(* Logix 5000 project; controller FV vendor 1 type 14 code 217 rev 31.11; software revision 31.00; part 29 of 63 *)
(* tags used below, declared in another part *)
   Alarm_Reset : BOOL;
   Default_Check_Time : DINT;
   FR_FV30_AV01 : PlantItem;   // FV30_AV01
   FR_FV30_AV01_ALARM : ALARM_DIGITAL;
   FR_FV30_AV01_C : ALIAS FOR RIO_Rack_2:10:I.Data.4;
   FR_FV30_AV01_O : ALIAS FOR RIO_Rack_2:10:I.Data.0;
   FR_FV30_AV01_RDR : ALIAS FOR RIO_Rack_2:11:O.Data.0;
   FR_FV30_AV04 : PlantItem;   // FV30_AV04
   FR_FV30_AV04_ALARM : ALARM_DIGITAL;
   FR_FV30_AV04_C : ALIAS FOR RIO_Rack_2:10:I.Data.5;
   FR_FV30_AV04_DR : ALIAS FOR RIO_Rack_2:11:O.Data.1;
   FR_FV30_AV04_O : ALIAS FOR RIO_Rack_2:10:I.Data.1;
   FR_FV30_AV05 : PlantItem;   // FV30_AV05
   FR_FV30_AV05_ALARM : ALARM_DIGITAL;
   FR_FV30_AV05_C : ALIAS FOR RIO_Rack_2:10:I.Data.6;
   FR_FV30_AV05_DR : ALIAS FOR RIO_Rack_2:11:O.Data.2;
   FR_FV30_AV05_O : ALIAS FOR RIO_Rack_2:10:I.Data.2;
   FR_FV30_AV06 : PlantItem;   // FV30_AV06
   FR_FV30_AV06_ALARM : ALARM_DIGITAL;
   FR_FV30_AV06_C : ALIAS FOR RIO_Rack_2:10:I.Data.7;
   FR_FV30_AV06_DR : ALIAS FOR RIO_Rack_2:11:O.Data.3;
   FR_FV30_AV06_O : ALIAS FOR RIO_Rack_2:10:I.Data.3;
   FR_FV30_AV07 : PlantItem;   // FV30_AV07
   FR_FV30_AV07_ALARM : ALARM_DIGITAL;
   FR_FV30_AV07_C : ALIAS FOR RIO_Rack_2:10:I.Data.12;
   FR_FV30_AV07_DR : ALIAS FOR RIO_Rack_2:11:O.Data.4;
   FR_FV30_AV07_O : ALIAS FOR RIO_Rack_2:10:I.Data.8;
   FR_VB4_AV04 : PlantItem;   // VB4_AV04
   FR_VB4_AV04_ALARM : ALARM_DIGITAL;
   FR_VB4_AV04_C : ALIAS FOR RIO_Rack_2:7:I.Data.29;
   FR_VB4_AV04_DR : ALIAS FOR RIO_Rack_2:8:O.Data.13;
   FR_VB4_AV04_O : ALIAS FOR RIO_Rack_2:7:I.Data.25;
   FR_VB4_AV05 : PlantItem;   // VB4_AV05
   FR_VB4_AV05_ALARM : ALARM_DIGITAL;
   FR_VB4_AV05_C : ALIAS FOR RIO_Rack_2:7:I.Data.30;
   FR_VB4_AV05_DR : ALIAS FOR RIO_Rack_2:8:O.Data.14;
   FR_VB4_AV05_O : ALIAS FOR RIO_Rack_2:7:I.Data.26;
   FR_VB4_AV06 : PlantItem;   // VB4_AV06
   FR_VB4_AV06_ALARM : ALARM_DIGITAL;
   FR_VB4_AV06_C : ALIAS FOR RIO_Rack_2:7:I.Data.31;
   FR_VB4_AV06_DR : ALIAS FOR RIO_Rack_2:8:O.Data.15;
   FR_VB4_AV06_O : ALIAS FOR RIO_Rack_2:7:I.Data.27;
   FR_VB4_AV07 : PlantItem;   // VB4_AV07
   FR_VB4_AV07_ALARM : ALARM_DIGITAL;
   FR_VB4_AV07_C : ALIAS FOR RIO_Rack_2:9:I.Data.4;
   FR_VB4_AV07_DR : ALIAS FOR RIO_Rack_2:8:O.Data.16;
   FR_VB4_AV07_O : ALIAS FOR RIO_Rack_2:9:I.Data.0;
   FR_VB4_AV08 : PlantItem;   // VB4_AV08
   FR_VB4_AV08_ALARM : ALARM_DIGITAL;
   FR_VB4_AV08_C : ALIAS FOR RIO_Rack_2:9:I.Data.5;
   FR_VB4_AV08_DR : ALIAS FOR RIO_Rack_2:8:O.Data.17;
   FR_VB4_AV08_O : ALIAS FOR RIO_Rack_2:9:I.Data.1;
   FR_VB4_AV09 : PlantItem;   // VB4_AV09
   FR_VB4_AV09_ALARM : ALARM_DIGITAL;
   FR_VB4_AV09_C : ALIAS FOR RIO_Rack_2:9:I.Data.6;
   FR_VB4_AV09_DR : ALIAS FOR RIO_Rack_2:8:O.Data.18;
   FR_VB4_AV09_O : ALIAS FOR RIO_Rack_2:9:I.Data.2;
   FR_VB4_AV10 : PlantItem;   // VB4_AV10
   FR_VB4_AV10_ALARM : ALARM_DIGITAL;
   FR_VB4_AV10_C : ALIAS FOR RIO_Rack_2:9:I.Data.7;
   FR_VB4_AV10_DR : ALIAS FOR RIO_Rack_2:8:O.Data.19;
   FR_VB4_AV10_O : ALIAS FOR RIO_Rack_2:9:I.Data.3;
   FR_VB4_AV11 : PlantItem;   // VB4_AV11
   FR_VB4_AV11_ALARM : ALARM_DIGITAL;
   FR_VB4_AV11_C : ALIAS FOR RIO_Rack_2:9:I.Data.12;
   FR_VB4_AV11_DR : ALIAS FOR RIO_Rack_2:8:O.Data.20;
   FR_VB4_AV11_O : ALIAS FOR RIO_Rack_2:9:I.Data.8;
   FR_VB4_AV12 : PlantItem;   // VB4_AV12
   FR_VB4_AV12_ALARM : ALARM_DIGITAL;
   FR_VB4_AV12_C : ALIAS FOR RIO_Rack_2:9:I.Data.13;
   FR_VB4_AV12_DR : ALIAS FOR RIO_Rack_2:8:O.Data.21;
   FR_VB4_AV12_O : ALIAS FOR RIO_Rack_2:9:I.Data.9;
   FR_VB4_AV13 : PlantItem;   // VB4_AV13
   FR_VB4_AV13_ALARM : ALARM_DIGITAL;
   FR_VB4_AV13_C : ALIAS FOR RIO_Rack_2:9:I.Data.14;
   FR_VB4_AV13_DR : ALIAS FOR RIO_Rack_2:8:O.Data.22;
   FR_VB4_AV13_O : ALIAS FOR RIO_Rack_2:9:I.Data.10;
   FR_VB4_AV14 : PlantItem;   // VB4_AV14
   FR_VB4_AV14_ALARM : ALARM_DIGITAL;
   FR_VB4_AV14_C : ALIAS FOR RIO_Rack_2:9:I.Data.15;
   FR_VB4_AV14_DR : ALIAS FOR RIO_Rack_2:8:O.Data.23;
   FR_VB4_AV14_O : ALIAS FOR RIO_Rack_2:9:I.Data.11;
   FR_VB4_AV15 : PlantItem;   // VB4_AV15
   FR_VB4_AV15_ALARM : ALARM_DIGITAL;
   FR_VB4_AV15_C : ALIAS FOR RIO_Rack_2:9:I.Data.20;
   FR_VB4_AV15_DR : ALIAS FOR RIO_Rack_2:8:O.Data.24;
   FR_VB4_AV15_O : ALIAS FOR RIO_Rack_2:9:I.Data.16;
   FR_VB4_AV17 : PlantItem;   // VB4_AV17
   FR_VB4_AV17_ALARM : ALARM_DIGITAL;
   FR_VB4_AV17_C : ALIAS FOR RIO_Rack_2:9:I.Data.22;
   FR_VB4_AV17_DR : ALIAS FOR RIO_Rack_2:8:O.Data.26;
   FR_VB4_AV17_O : ALIAS FOR RIO_Rack_2:9:I.Data.18;
   FR_VB4_AV18 : PlantItem;   // VB4_AV18
   FR_VB4_AV18_ALARM : ALARM_DIGITAL;
   FR_VB4_AV18_C : ALIAS FOR RIO_Rack_2:9:I.Data.23;
   FR_VB4_AV18_DR : ALIAS FOR RIO_Rack_2:8:O.Data.27;
   FR_VB4_AV18_O : ALIAS FOR RIO_Rack_2:9:I.Data.19;
   FR_VB4_AV19 : PlantItem;   // VB4_AV19
   FR_VB4_AV19_ALARM : ALARM_DIGITAL;
   FR_VB4_AV19_C : ALIAS FOR RIO_Rack_2:9:I.Data.28;
   FR_VB4_AV19_DR : ALIAS FOR RIO_Rack_2:8:O.Data.28;
   FR_VB4_AV19_O : ALIAS FOR RIO_Rack_2:9:I.Data.24;
   FR_VB4_AV20 : PlantItem;   // VB4_AV20
   FR_VB4_AV20_ALARM : ALARM_DIGITAL;
   FR_VB4_AV20_C : ALIAS FOR RIO_Rack_2:9:I.Data.29;
   FR_VB4_AV20_DR : ALIAS FOR RIO_Rack_2:8:O.Data.29;
   FR_VB4_AV20_O : ALIAS FOR RIO_Rack_2:9:I.Data.25;
   FR_VB4_AV21 : PlantItem;   // VB4_AV21
   FR_VB4_AV21_ALARM : ALARM_DIGITAL;
   FR_VB4_AV21_C : ALIAS FOR RIO_Rack_2:9:I.Data.30;
   FR_VB4_AV21_DR : ALIAS FOR RIO_Rack_2:8:O.Data.30;
   FR_VB4_AV21_O : ALIAS FOR RIO_Rack_2:9:I.Data.26;
   FR_VB4_AV22 : PlantItem;   // VB4_AV22
   FR_VB4_AV22_ALARM : ALARM_DIGITAL;
   FR_VB4_AV22_C : ALIAS FOR RIO_Rack_2:9:I.Data.31;
   FR_VB4_AV22_DR : ALIAS FOR RIO_Rack_2:8:O.Data.31;
   FR_VB4_AV22_O : ALIAS FOR RIO_Rack_2:9:I.Data.27;
   FR_VB4_AV23 : PlantItem;   // VB4_AV23
   FR_VB4_AV23_ALARM : ALARM_DIGITAL;
   FR_VB4_AV23_C : ALIAS FOR RIO_Rack_2:9:I.Data.21;
   FR_VB4_AV23_DR : ALIAS FOR RIO_Rack_2:8:O.Data.25;
   FR_VB4_AV23_O : ALIAS FOR RIO_Rack_2:9:I.Data.17;
   Item_Faults_Are_Latched : BOOL;
   Item_Simulation_Flag : BOOL;
   One_Second_One_Scan : ALIAS FOR One_Second_1_scan;
(* FR_Common, continued *)

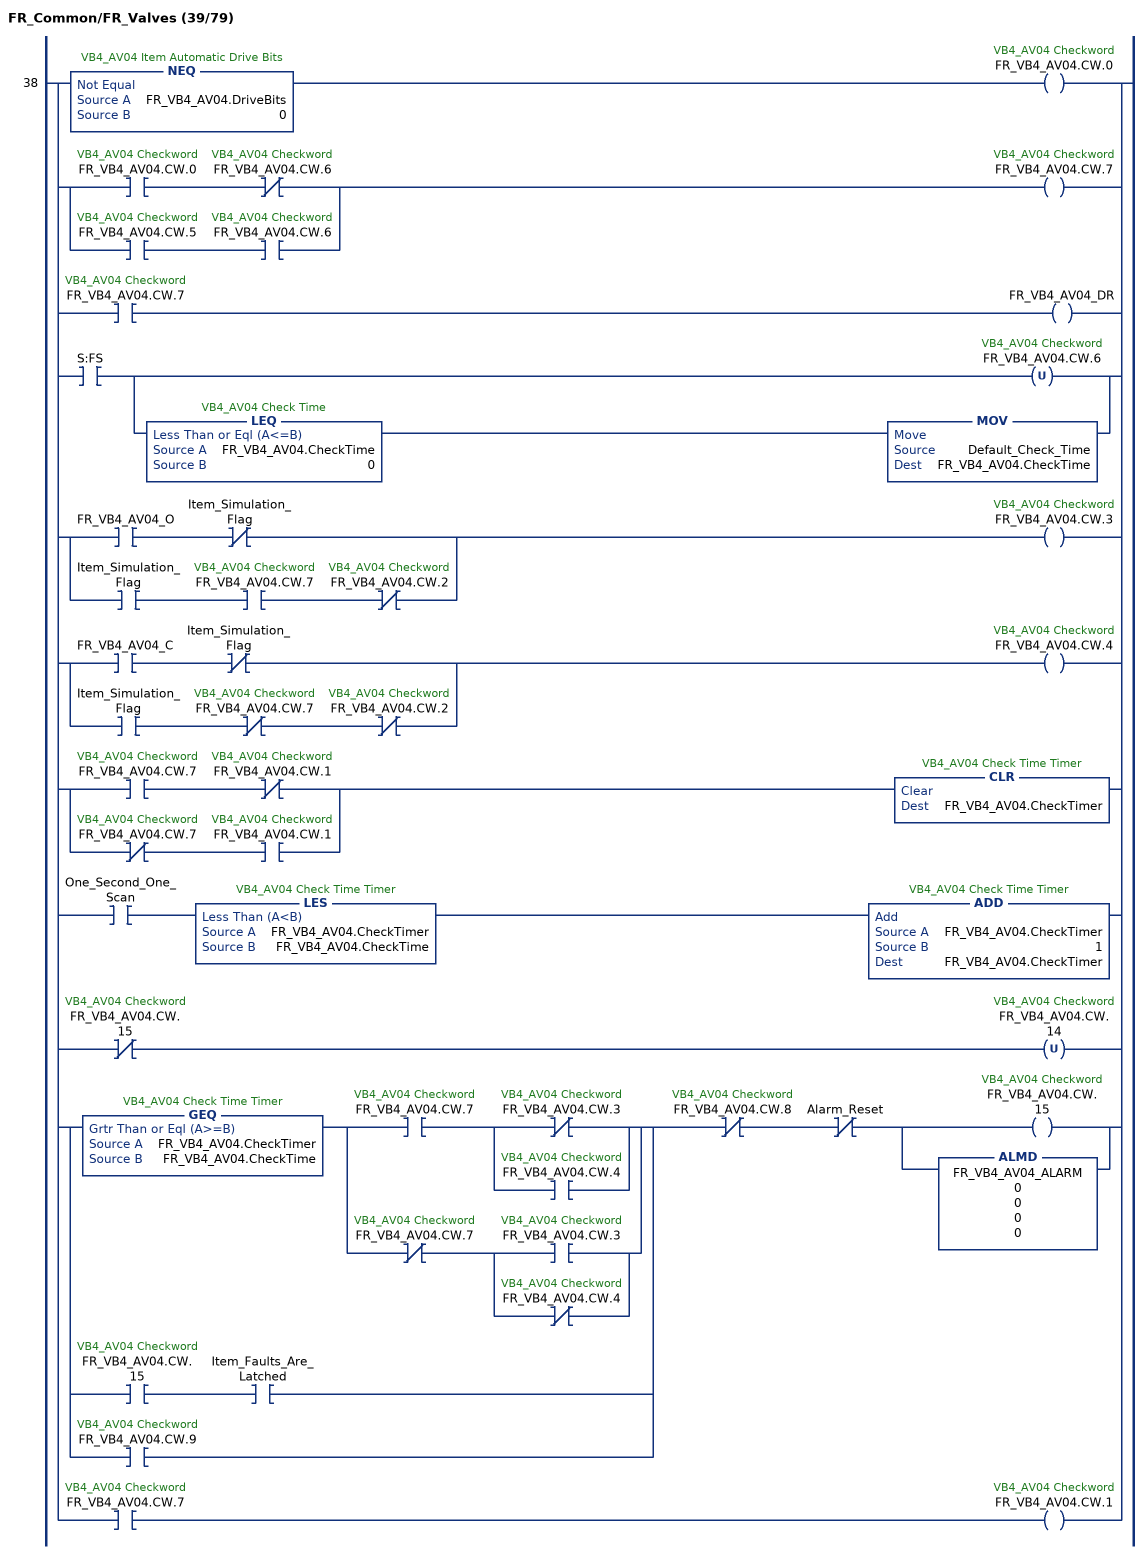
   [picture p592: FR_Common/FR_Valves rungs 38-38]
   38: [NEQ(FR_VB4_AV04.DriveBits,0) OTE(FR_VB4_AV04.CW.0) ,[XIC(FR_VB4_AV04.CW.0) XIO(FR_VB4_AV04.CW.6) ,XIC(FR_VB4_AV04.CW.5) XIC(FR_VB4_AV04.CW.6) ] OTE(FR_VB4_AV04.CW.7) ,XIC(FR_VB4_AV04.CW.7) OTE(FR_VB4_AV04_DR) ,XIC(S:FS) [OTU(FR_VB4_AV04.CW.6) ,LEQ(FR_VB4_AV04.CheckTime,0) MOV(Default_Check_Time,FR_VB4_AV04.CheckTime) ] ,[[XIC(FR_VB4_AV04_O) XIO(Item_Simulation_Flag) ,XIC(Item_Simulation_Flag) XIC(FR_VB4_AV04.CW.7) XIO(FR_VB4_AV04.CW.2) ] OTE(FR_VB4_AV04.CW.3) ,[XIC(FR_VB4_AV04_C) XIO(Item_Simulation_Flag) ,XIC(Item_Simulation_Flag) XIO(FR_VB4_AV04.CW.7) XIO(FR_VB4_AV04.CW.2) ] OTE(FR_VB4_AV04.CW.4) ] ,[XIC(FR_VB4_AV04.CW.7) XIO(FR_VB4_AV04.CW.1) ,XIO(FR_VB4_AV04.CW.7) XIC(FR_VB4_AV04.CW.1) ] CLR(FR_VB4_AV04.CheckTimer) ,XIC(One_Second_One_Scan) LES(FR_VB4_AV04.CheckTimer,FR_VB4_AV04.CheckTime) ADD(FR_VB4_AV04.CheckTimer,1,FR_VB4_AV04.CheckTimer) ,XIO(FR_VB4_AV04.CW.15) OTU(FR_VB4_AV04.CW.14) ,[GEQ(FR_VB4_AV04.CheckTimer,FR_VB4_AV04.CheckTime) [XIC(FR_VB4_AV04.CW.7) [XIO(FR_VB4_AV04.CW.3) ,XIC(FR_VB4_AV04.CW.4) ] ,XIO(FR_VB4_AV04.CW.7) [XIC(FR_VB4_AV04.CW.3) ,XIO(FR_VB4_AV04.CW.4) ] ] ,XIC(FR_VB4_AV04.CW.15) XIC(Item_Faults_Are_Latched) ,XIC(FR_VB4_AV04.CW.9) ] XIO(FR_VB4_AV04.CW.8) XIO(Alarm_Reset) [OTE(FR_VB4_AV04.CW.15) ,ALMD(FR_VB4_AV04_ALARM,0,0,0,0) ] ,XIC(FR_VB4_AV04.CW.7) OTE(FR_VB4_AV04.CW.1) ];
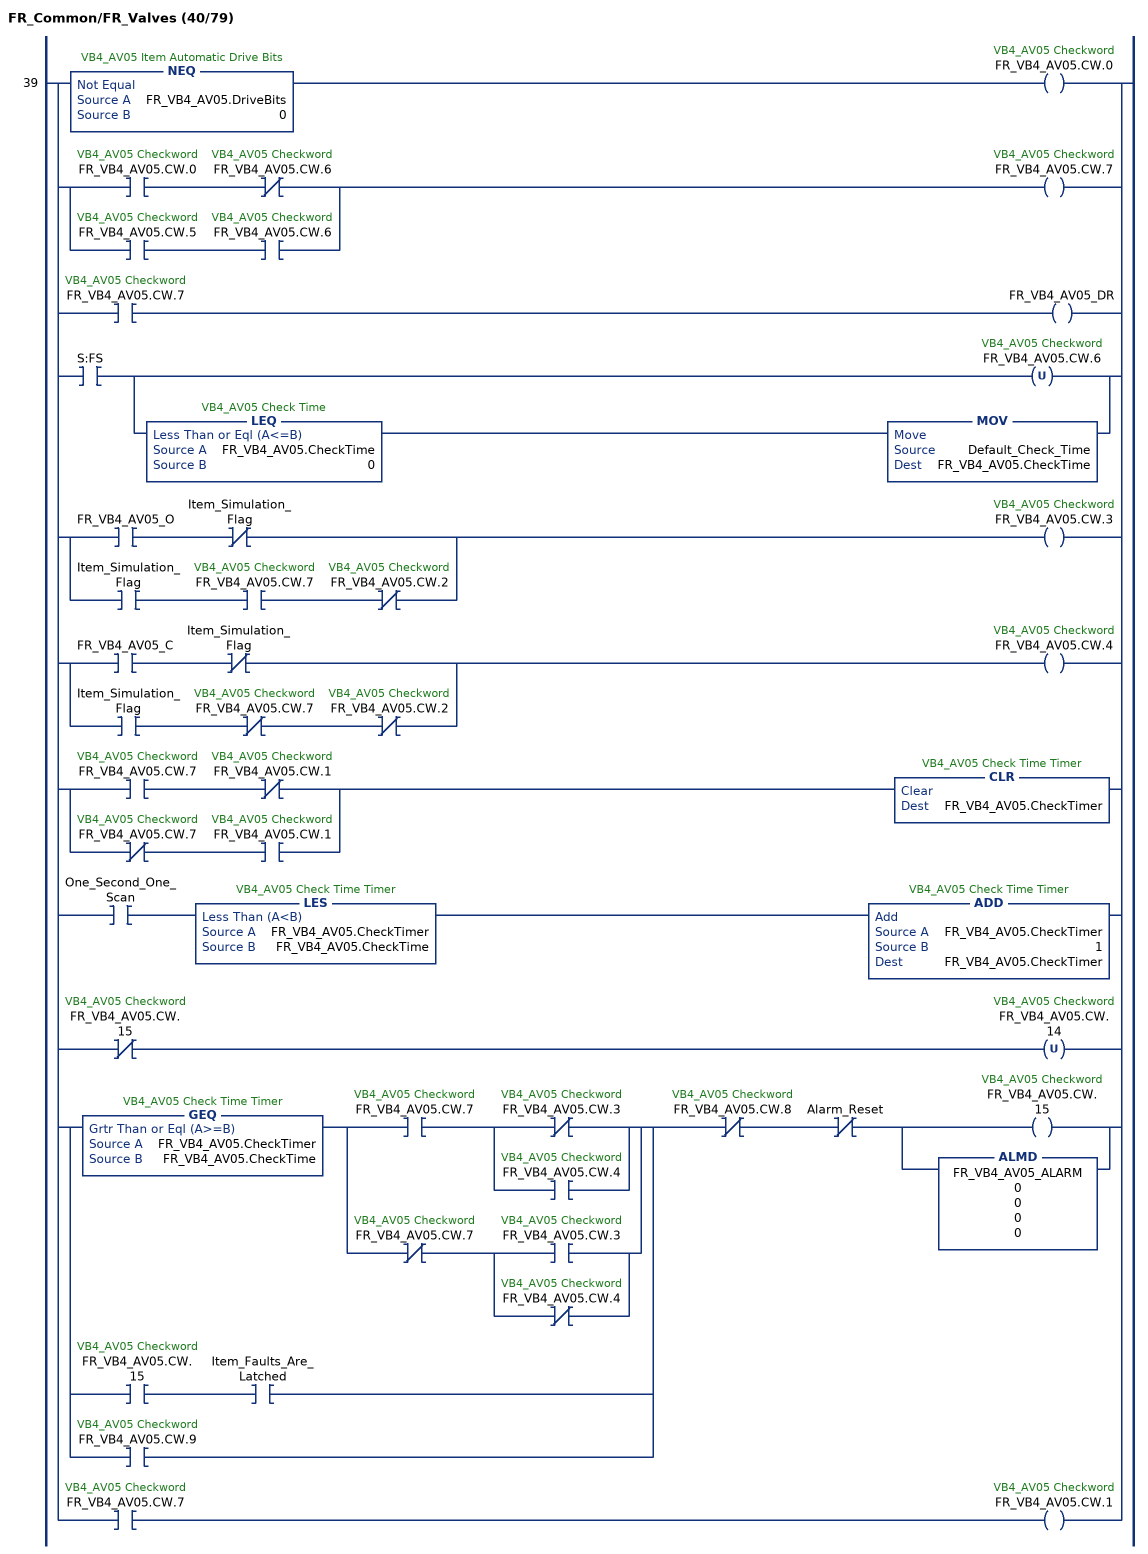
   39: [NEQ(FR_VB4_AV05.DriveBits,0) OTE(FR_VB4_AV05.CW.0) ,[XIC(FR_VB4_AV05.CW.0) XIO(FR_VB4_AV05.CW.6) ,XIC(FR_VB4_AV05.CW.5) XIC(FR_VB4_AV05.CW.6) ] OTE(FR_VB4_AV05.CW.7) ,XIC(FR_VB4_AV05.CW.7) OTE(FR_VB4_AV05_DR) ,XIC(S:FS) [OTU(FR_VB4_AV05.CW.6) ,LEQ(FR_VB4_AV05.CheckTime,0) MOV(Default_Check_Time,FR_VB4_AV05.CheckTime) ] ,[[XIC(FR_VB4_AV05_O) XIO(Item_Simulation_Flag) ,XIC(Item_Simulation_Flag) XIC(FR_VB4_AV05.CW.7) XIO(FR_VB4_AV05.CW.2) ] OTE(FR_VB4_AV05.CW.3) ,[XIC(FR_VB4_AV05_C) XIO(Item_Simulation_Flag) ,XIC(Item_Simulation_Flag) XIO(FR_VB4_AV05.CW.7) XIO(FR_VB4_AV05.CW.2) ] OTE(FR_VB4_AV05.CW.4) ] ,[XIC(FR_VB4_AV05.CW.7) XIO(FR_VB4_AV05.CW.1) ,XIO(FR_VB4_AV05.CW.7) XIC(FR_VB4_AV05.CW.1) ] CLR(FR_VB4_AV05.CheckTimer) ,XIC(One_Second_One_Scan) LES(FR_VB4_AV05.CheckTimer,FR_VB4_AV05.CheckTime) ADD(FR_VB4_AV05.CheckTimer,1,FR_VB4_AV05.CheckTimer) ,XIO(FR_VB4_AV05.CW.15) OTU(FR_VB4_AV05.CW.14) ,[GEQ(FR_VB4_AV05.CheckTimer,FR_VB4_AV05.CheckTime) [XIC(FR_VB4_AV05.CW.7) [XIO(FR_VB4_AV05.CW.3) ,XIC(FR_VB4_AV05.CW.4) ] ,XIO(FR_VB4_AV05.CW.7) [XIC(FR_VB4_AV05.CW.3) ,XIO(FR_VB4_AV05.CW.4) ] ] ,XIC(FR_VB4_AV05.CW.15) XIC(Item_Faults_Are_Latched) ,XIC(FR_VB4_AV05.CW.9) ] XIO(FR_VB4_AV05.CW.8) XIO(Alarm_Reset) [OTE(FR_VB4_AV05.CW.15) ,ALMD(FR_VB4_AV05_ALARM,0,0,0,0) ] ,XIC(FR_VB4_AV05.CW.7) OTE(FR_VB4_AV05.CW.1) ];
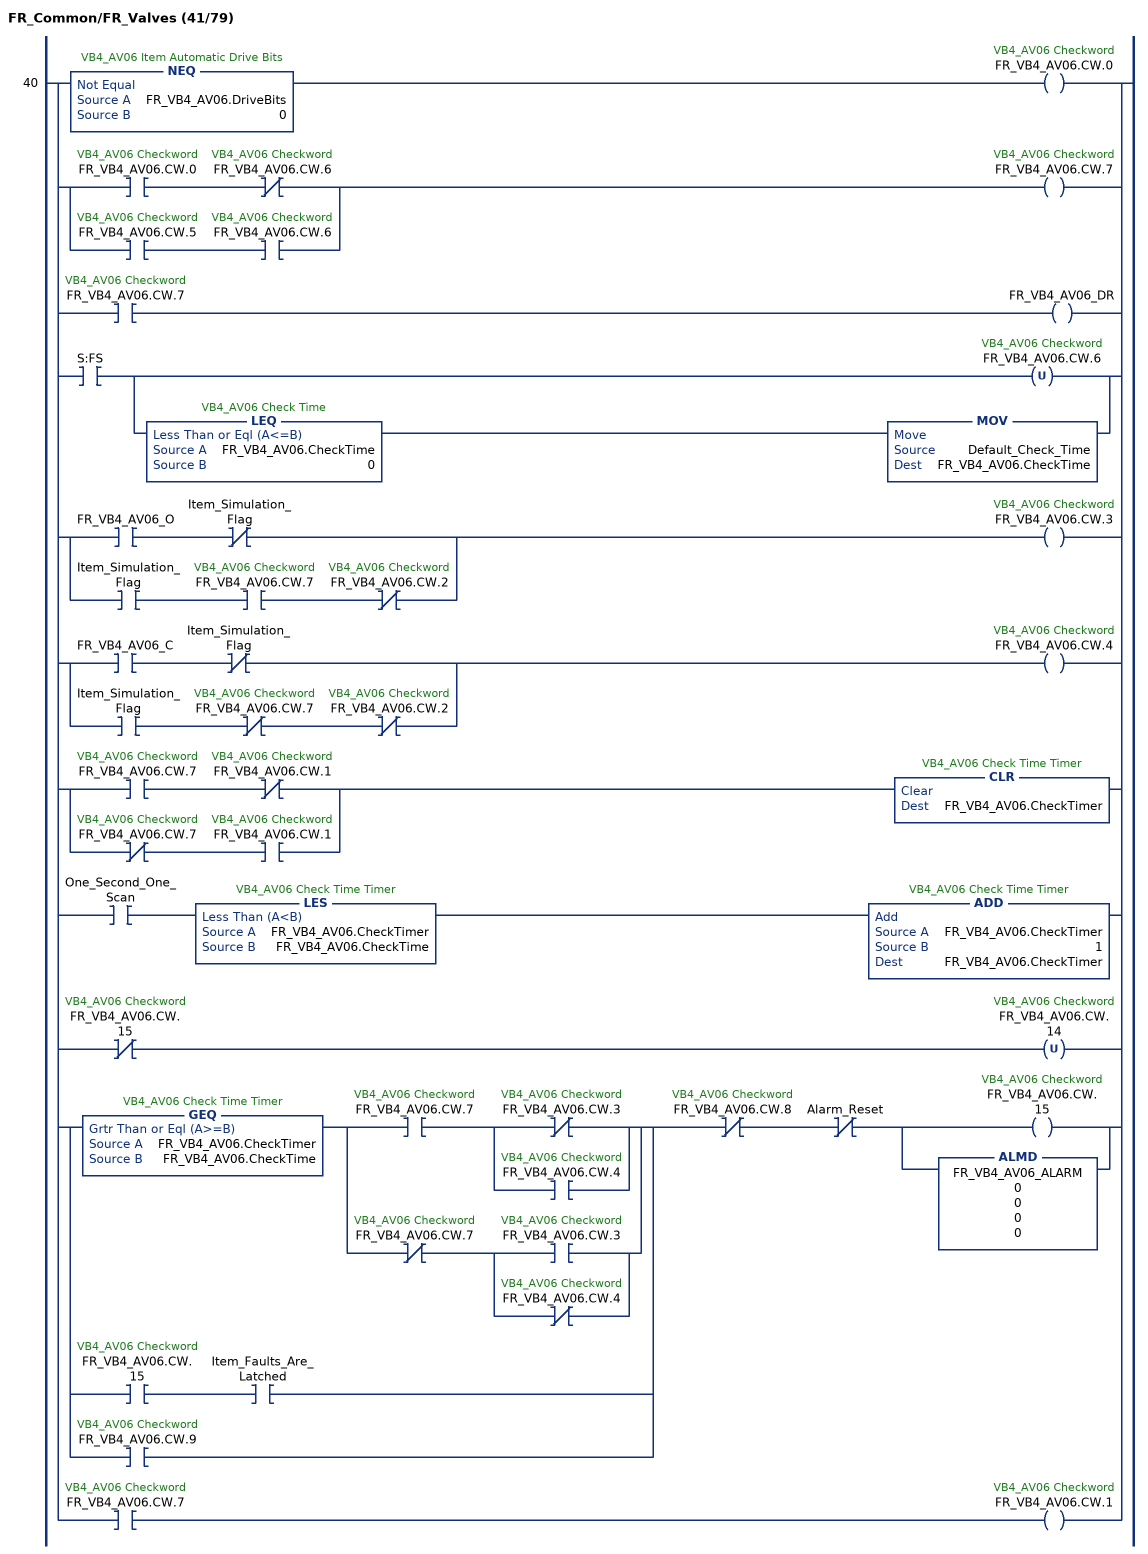
   40: [NEQ(FR_VB4_AV06.DriveBits,0) OTE(FR_VB4_AV06.CW.0) ,[XIC(FR_VB4_AV06.CW.0) XIO(FR_VB4_AV06.CW.6) ,XIC(FR_VB4_AV06.CW.5) XIC(FR_VB4_AV06.CW.6) ] OTE(FR_VB4_AV06.CW.7) ,XIC(FR_VB4_AV06.CW.7) OTE(FR_VB4_AV06_DR) ,XIC(S:FS) [OTU(FR_VB4_AV06.CW.6) ,LEQ(FR_VB4_AV06.CheckTime,0) MOV(Default_Check_Time,FR_VB4_AV06.CheckTime) ] ,[[XIC(FR_VB4_AV06_O) XIO(Item_Simulation_Flag) ,XIC(Item_Simulation_Flag) XIC(FR_VB4_AV06.CW.7) XIO(FR_VB4_AV06.CW.2) ] OTE(FR_VB4_AV06.CW.3) ,[XIC(FR_VB4_AV06_C) XIO(Item_Simulation_Flag) ,XIC(Item_Simulation_Flag) XIO(FR_VB4_AV06.CW.7) XIO(FR_VB4_AV06.CW.2) ] OTE(FR_VB4_AV06.CW.4) ] ,[XIC(FR_VB4_AV06.CW.7) XIO(FR_VB4_AV06.CW.1) ,XIO(FR_VB4_AV06.CW.7) XIC(FR_VB4_AV06.CW.1) ] CLR(FR_VB4_AV06.CheckTimer) ,XIC(One_Second_One_Scan) LES(FR_VB4_AV06.CheckTimer,FR_VB4_AV06.CheckTime) ADD(FR_VB4_AV06.CheckTimer,1,FR_VB4_AV06.CheckTimer) ,XIO(FR_VB4_AV06.CW.15) OTU(FR_VB4_AV06.CW.14) ,[GEQ(FR_VB4_AV06.CheckTimer,FR_VB4_AV06.CheckTime) [XIC(FR_VB4_AV06.CW.7) [XIO(FR_VB4_AV06.CW.3) ,XIC(FR_VB4_AV06.CW.4) ] ,XIO(FR_VB4_AV06.CW.7) [XIC(FR_VB4_AV06.CW.3) ,XIO(FR_VB4_AV06.CW.4) ] ] ,XIC(FR_VB4_AV06.CW.15) XIC(Item_Faults_Are_Latched) ,XIC(FR_VB4_AV06.CW.9) ] XIO(FR_VB4_AV06.CW.8) XIO(Alarm_Reset) [OTE(FR_VB4_AV06.CW.15) ,ALMD(FR_VB4_AV06_ALARM,0,0,0,0) ] ,XIC(FR_VB4_AV06.CW.7) OTE(FR_VB4_AV06.CW.1) ];
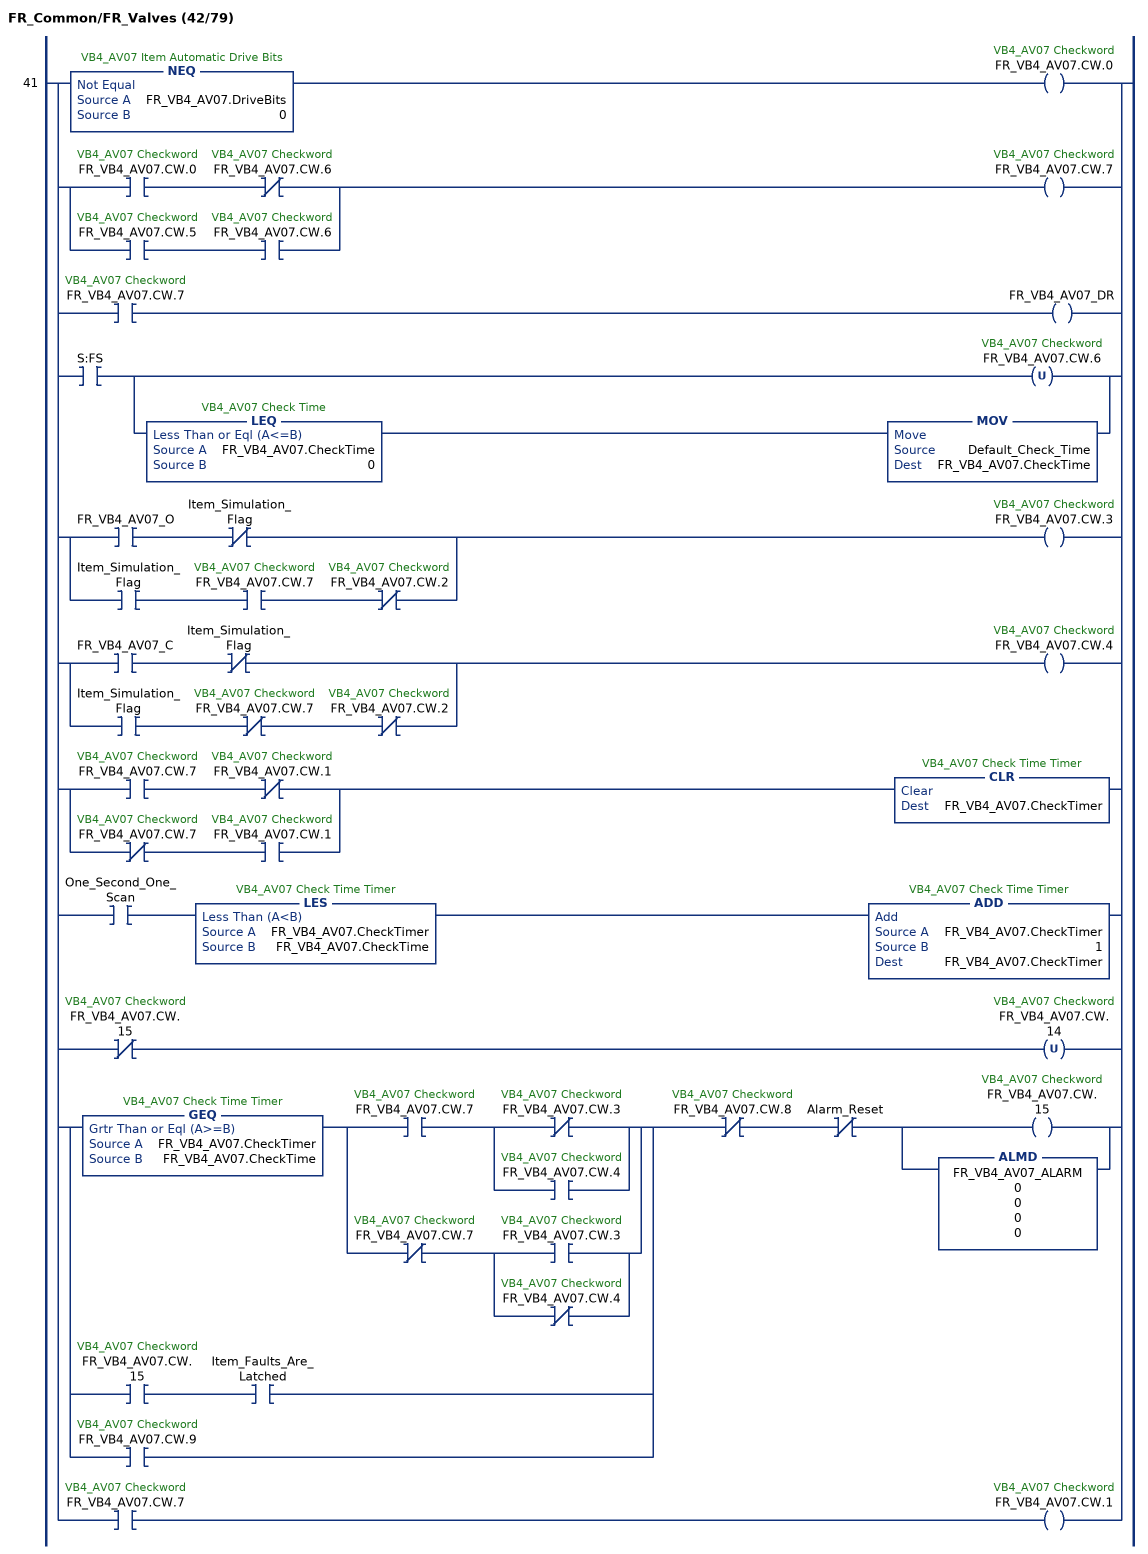
   41: [NEQ(FR_VB4_AV07.DriveBits,0) OTE(FR_VB4_AV07.CW.0) ,[XIC(FR_VB4_AV07.CW.0) XIO(FR_VB4_AV07.CW.6) ,XIC(FR_VB4_AV07.CW.5) XIC(FR_VB4_AV07.CW.6) ] OTE(FR_VB4_AV07.CW.7) ,XIC(FR_VB4_AV07.CW.7) OTE(FR_VB4_AV07_DR) ,XIC(S:FS) [OTU(FR_VB4_AV07.CW.6) ,LEQ(FR_VB4_AV07.CheckTime,0) MOV(Default_Check_Time,FR_VB4_AV07.CheckTime) ] ,[[XIC(FR_VB4_AV07_O) XIO(Item_Simulation_Flag) ,XIC(Item_Simulation_Flag) XIC(FR_VB4_AV07.CW.7) XIO(FR_VB4_AV07.CW.2) ] OTE(FR_VB4_AV07.CW.3) ,[XIC(FR_VB4_AV07_C) XIO(Item_Simulation_Flag) ,XIC(Item_Simulation_Flag) XIO(FR_VB4_AV07.CW.7) XIO(FR_VB4_AV07.CW.2) ] OTE(FR_VB4_AV07.CW.4) ] ,[XIC(FR_VB4_AV07.CW.7) XIO(FR_VB4_AV07.CW.1) ,XIO(FR_VB4_AV07.CW.7) XIC(FR_VB4_AV07.CW.1) ] CLR(FR_VB4_AV07.CheckTimer) ,XIC(One_Second_One_Scan) LES(FR_VB4_AV07.CheckTimer,FR_VB4_AV07.CheckTime) ADD(FR_VB4_AV07.CheckTimer,1,FR_VB4_AV07.CheckTimer) ,XIO(FR_VB4_AV07.CW.15) OTU(FR_VB4_AV07.CW.14) ,[GEQ(FR_VB4_AV07.CheckTimer,FR_VB4_AV07.CheckTime) [XIC(FR_VB4_AV07.CW.7) [XIO(FR_VB4_AV07.CW.3) ,XIC(FR_VB4_AV07.CW.4) ] ,XIO(FR_VB4_AV07.CW.7) [XIC(FR_VB4_AV07.CW.3) ,XIO(FR_VB4_AV07.CW.4) ] ] ,XIC(FR_VB4_AV07.CW.15) XIC(Item_Faults_Are_Latched) ,XIC(FR_VB4_AV07.CW.9) ] XIO(FR_VB4_AV07.CW.8) XIO(Alarm_Reset) [OTE(FR_VB4_AV07.CW.15) ,ALMD(FR_VB4_AV07_ALARM,0,0,0,0) ] ,XIC(FR_VB4_AV07.CW.7) OTE(FR_VB4_AV07.CW.1) ];
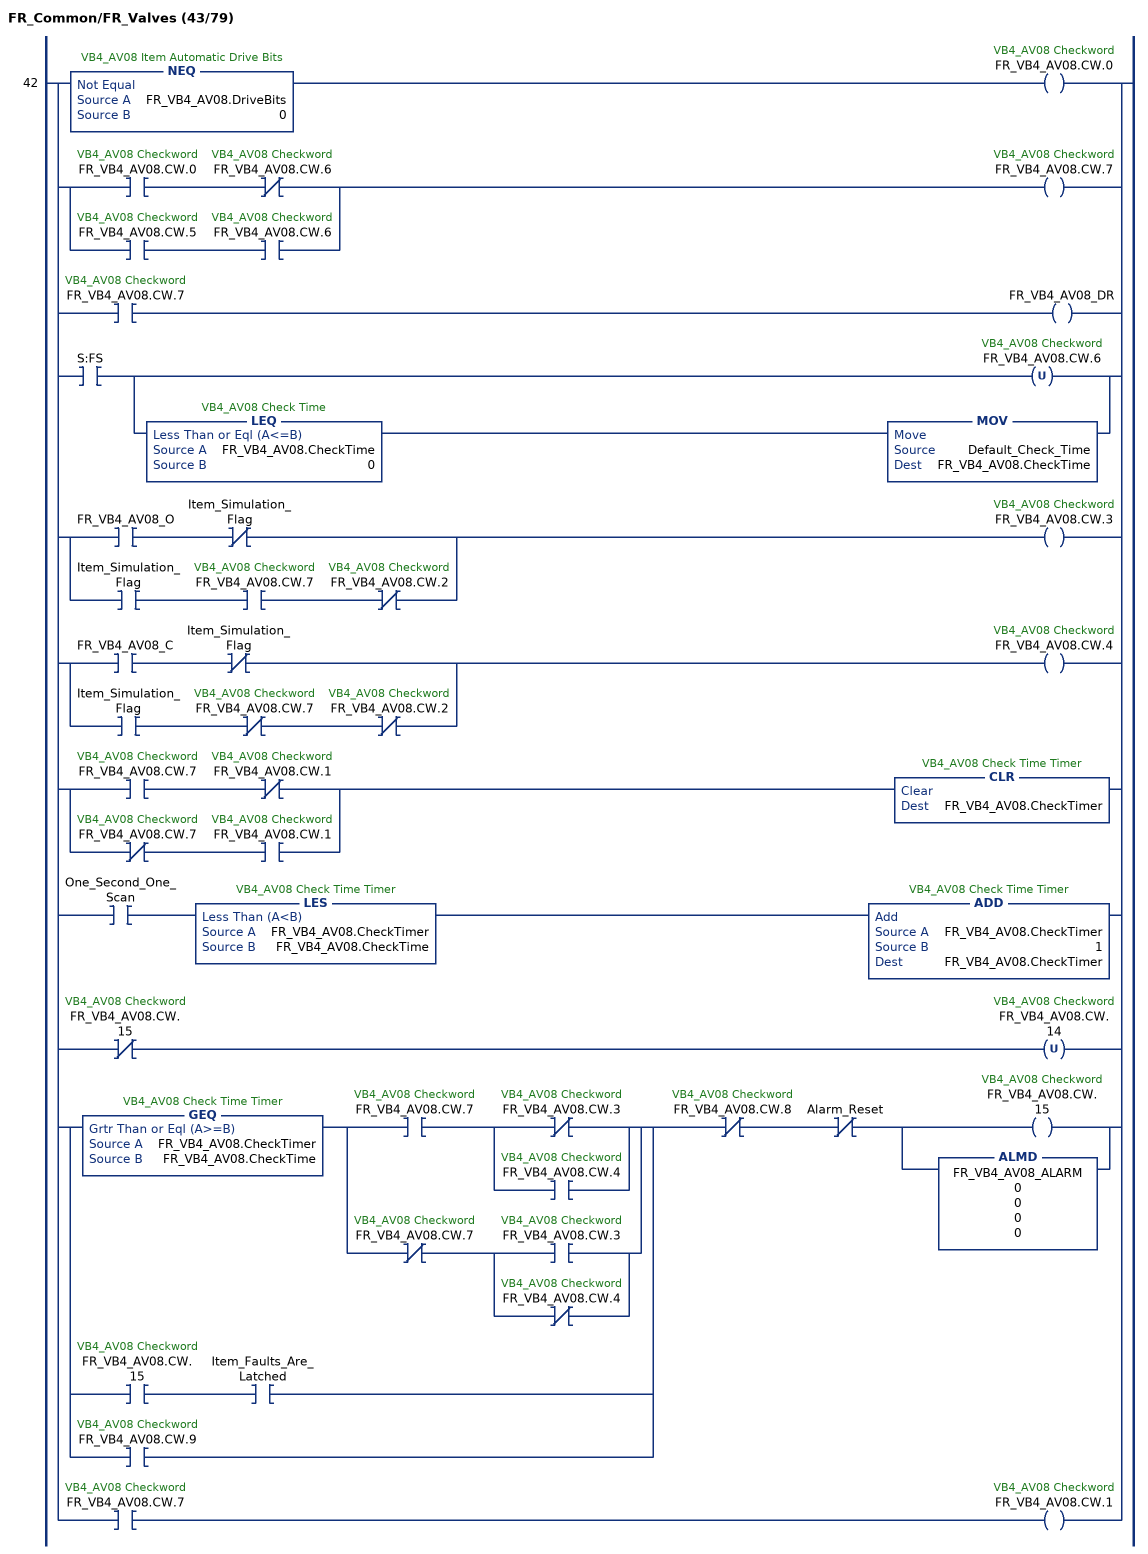
   42: [NEQ(FR_VB4_AV08.DriveBits,0) OTE(FR_VB4_AV08.CW.0) ,[XIC(FR_VB4_AV08.CW.0) XIO(FR_VB4_AV08.CW.6) ,XIC(FR_VB4_AV08.CW.5) XIC(FR_VB4_AV08.CW.6) ] OTE(FR_VB4_AV08.CW.7) ,XIC(FR_VB4_AV08.CW.7) OTE(FR_VB4_AV08_DR) ,XIC(S:FS) [OTU(FR_VB4_AV08.CW.6) ,LEQ(FR_VB4_AV08.CheckTime,0) MOV(Default_Check_Time,FR_VB4_AV08.CheckTime) ] ,[[XIC(FR_VB4_AV08_O) XIO(Item_Simulation_Flag) ,XIC(Item_Simulation_Flag) XIC(FR_VB4_AV08.CW.7) XIO(FR_VB4_AV08.CW.2) ] OTE(FR_VB4_AV08.CW.3) ,[XIC(FR_VB4_AV08_C) XIO(Item_Simulation_Flag) ,XIC(Item_Simulation_Flag) XIO(FR_VB4_AV08.CW.7) XIO(FR_VB4_AV08.CW.2) ] OTE(FR_VB4_AV08.CW.4) ] ,[XIC(FR_VB4_AV08.CW.7) XIO(FR_VB4_AV08.CW.1) ,XIO(FR_VB4_AV08.CW.7) XIC(FR_VB4_AV08.CW.1) ] CLR(FR_VB4_AV08.CheckTimer) ,XIC(One_Second_One_Scan) LES(FR_VB4_AV08.CheckTimer,FR_VB4_AV08.CheckTime) ADD(FR_VB4_AV08.CheckTimer,1,FR_VB4_AV08.CheckTimer) ,XIO(FR_VB4_AV08.CW.15) OTU(FR_VB4_AV08.CW.14) ,[GEQ(FR_VB4_AV08.CheckTimer,FR_VB4_AV08.CheckTime) [XIC(FR_VB4_AV08.CW.7) [XIO(FR_VB4_AV08.CW.3) ,XIC(FR_VB4_AV08.CW.4) ] ,XIO(FR_VB4_AV08.CW.7) [XIC(FR_VB4_AV08.CW.3) ,XIO(FR_VB4_AV08.CW.4) ] ] ,XIC(FR_VB4_AV08.CW.15) XIC(Item_Faults_Are_Latched) ,XIC(FR_VB4_AV08.CW.9) ] XIO(FR_VB4_AV08.CW.8) XIO(Alarm_Reset) [OTE(FR_VB4_AV08.CW.15) ,ALMD(FR_VB4_AV08_ALARM,0,0,0,0) ] ,XIC(FR_VB4_AV08.CW.7) OTE(FR_VB4_AV08.CW.1) ];
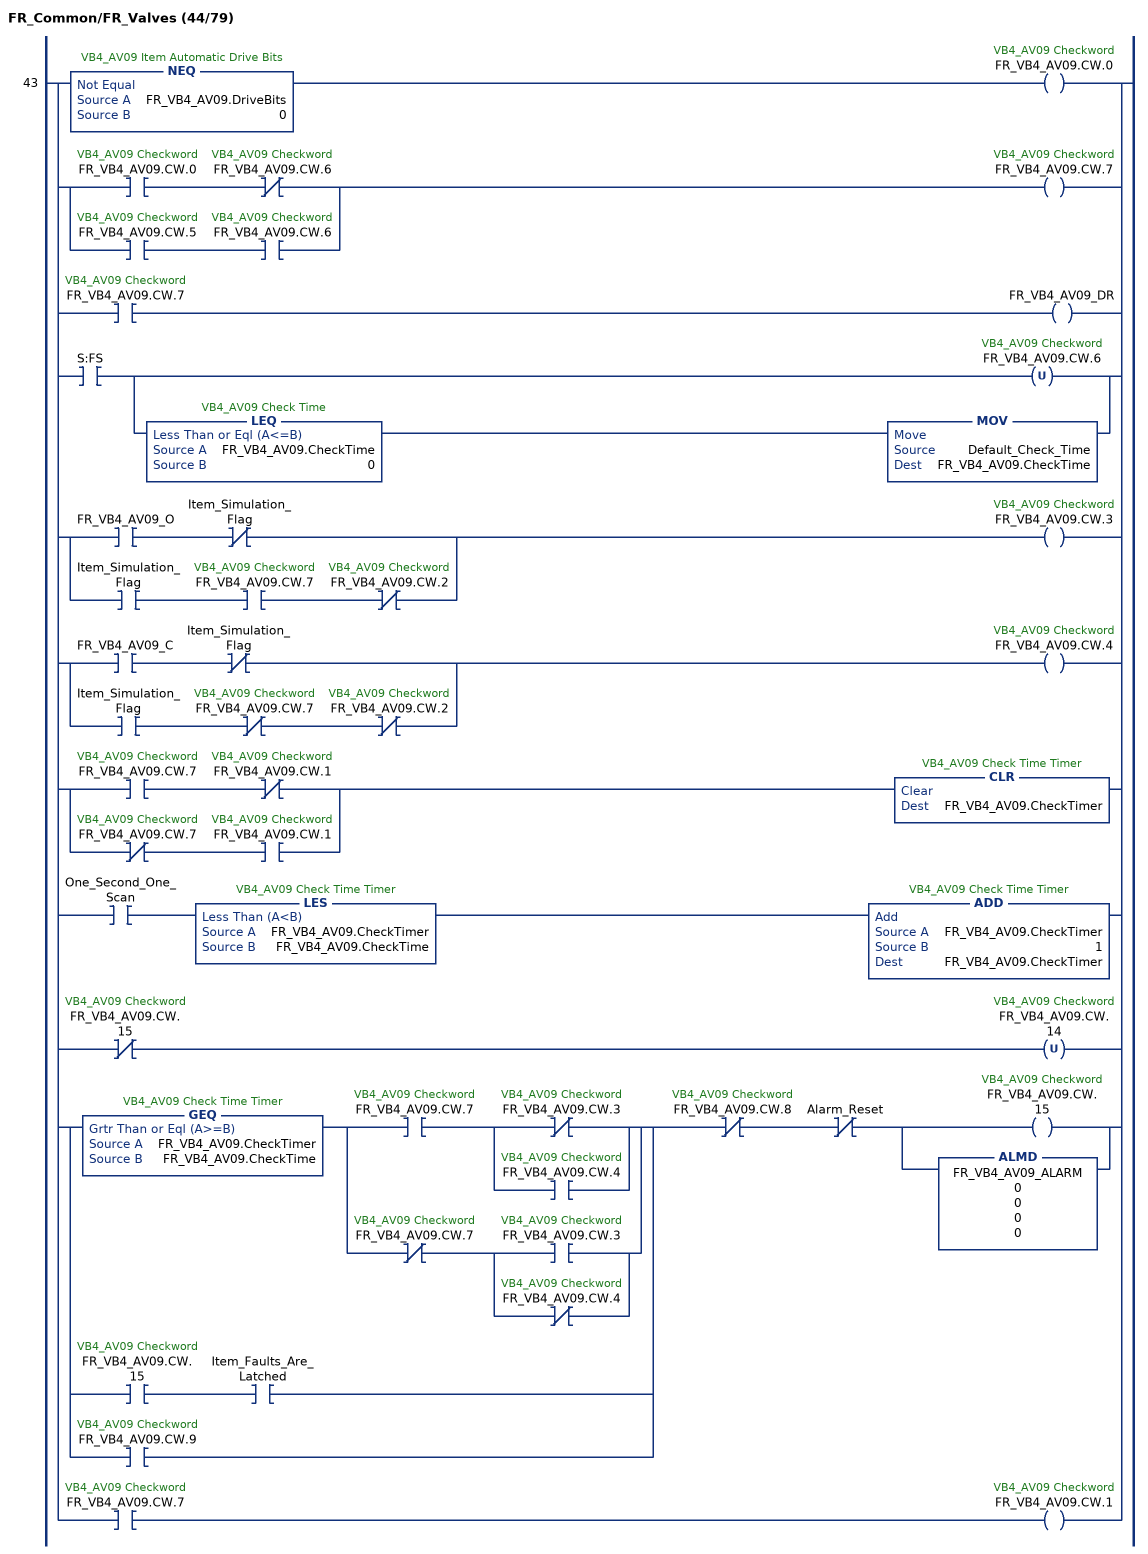
   43: [NEQ(FR_VB4_AV09.DriveBits,0) OTE(FR_VB4_AV09.CW.0) ,[XIC(FR_VB4_AV09.CW.0) XIO(FR_VB4_AV09.CW.6) ,XIC(FR_VB4_AV09.CW.5) XIC(FR_VB4_AV09.CW.6) ] OTE(FR_VB4_AV09.CW.7) ,XIC(FR_VB4_AV09.CW.7) OTE(FR_VB4_AV09_DR) ,XIC(S:FS) [OTU(FR_VB4_AV09.CW.6) ,LEQ(FR_VB4_AV09.CheckTime,0) MOV(Default_Check_Time,FR_VB4_AV09.CheckTime) ] ,[[XIC(FR_VB4_AV09_O) XIO(Item_Simulation_Flag) ,XIC(Item_Simulation_Flag) XIC(FR_VB4_AV09.CW.7) XIO(FR_VB4_AV09.CW.2) ] OTE(FR_VB4_AV09.CW.3) ,[XIC(FR_VB4_AV09_C) XIO(Item_Simulation_Flag) ,XIC(Item_Simulation_Flag) XIO(FR_VB4_AV09.CW.7) XIO(FR_VB4_AV09.CW.2) ] OTE(FR_VB4_AV09.CW.4) ] ,[XIC(FR_VB4_AV09.CW.7) XIO(FR_VB4_AV09.CW.1) ,XIO(FR_VB4_AV09.CW.7) XIC(FR_VB4_AV09.CW.1) ] CLR(FR_VB4_AV09.CheckTimer) ,XIC(One_Second_One_Scan) LES(FR_VB4_AV09.CheckTimer,FR_VB4_AV09.CheckTime) ADD(FR_VB4_AV09.CheckTimer,1,FR_VB4_AV09.CheckTimer) ,XIO(FR_VB4_AV09.CW.15) OTU(FR_VB4_AV09.CW.14) ,[GEQ(FR_VB4_AV09.CheckTimer,FR_VB4_AV09.CheckTime) [XIC(FR_VB4_AV09.CW.7) [XIO(FR_VB4_AV09.CW.3) ,XIC(FR_VB4_AV09.CW.4) ] ,XIO(FR_VB4_AV09.CW.7) [XIC(FR_VB4_AV09.CW.3) ,XIO(FR_VB4_AV09.CW.4) ] ] ,XIC(FR_VB4_AV09.CW.15) XIC(Item_Faults_Are_Latched) ,XIC(FR_VB4_AV09.CW.9) ] XIO(FR_VB4_AV09.CW.8) XIO(Alarm_Reset) [OTE(FR_VB4_AV09.CW.15) ,ALMD(FR_VB4_AV09_ALARM,0,0,0,0) ] ,XIC(FR_VB4_AV09.CW.7) OTE(FR_VB4_AV09.CW.1) ];